   PCmd_IntlkTripSuppress : ALIAS FOR IntlkTrip.PCmd_Suppress;   // Program Command to Suppress Interlock Trip Alarm
   PCmd_IntlkTripUnsuppress : ALIAS FOR IntlkTrip.PCmd_Unsuppress;   // Program Command to Unsuppress Interlock Trip Alarm
   PCmd_IntlkTripUnshelve : ALIAS FOR IntlkTrip.PCmd_Unshelve;   // Program Command to Unshelve Interlock Trip Alarm
   PCmd_IOFaultAck : ALIAS FOR IOFault.PCmd_Ack;   // Program Command to Acknowledge I/O Fault Alarm
   PCmd_IOFaultSuppress : ALIAS FOR IOFault.PCmd_Suppress;   // Program Command to Suppress I/O Fault Alarm
   PCmd_IOFaultUnsuppress : ALIAS FOR IOFault.PCmd_Unsuppress;   // Program Command to Unsuppress I/O Fault Alarm
   PCmd_IOFaultUnshelve : ALIAS FOR IOFault.PCmd_Unshelve;   // Program Command to Unshelve I/O Fault Alarm
   OCmd_Start : BOOL;   // Operator Command to Start Motor
   OCmd_Stop : BOOL;   // Operator Command to Stop Motor
   OCmd_Bypass : BOOL;   // Operator Command to Bypass all Bypassable Interlocks and Permissives
   OCmd_Check : BOOL;   // Operator Command to Check (not bypass) all Interlocks and Permissives
   MCmd_Disable : BOOL;   // Maintenance Command to Disable Motor
   MCmd_Enable : BOOL;   // Maintenance Command to Enable (allow to run) Motor
   OCmd_AcqLock : ALIAS FOR Mode.OCmd_AcqLock;
   OCmd_Unlock : ALIAS FOR Mode.OCmd_UnlockRel;
   OCmd_Reset : BOOL;   // Operator Command to Reset all Alarms requiring Reset
   OCmd_ResetAckAll : BOOL;   // Operator Command to Reset all Alarms and latched Shed conditions
END_VAR
VAR_OUTPUT
   Out_Run : BOOL; {access Read Only, visible}   // 1=Run Motor, 0=Stop Motor
   Out_Start : BOOL; {access Read Only, visible}   // 1=Start Motor, 0=Motor left in current state
   Out_Stop : BOOL; {access Read Only, visible}   // 1=Stop Motor, 0=Motor left in current state
   Val_Cmd : SINT; {access Read Only}   // Device Command 0=None, 1=Stop, 2=Start
   Val_Fdbk : SINT; {access Read Only}   // Device Feedback 0=Stopped, 1=Running
   Val_Sts : SINT; {access Read Only}   // Device Confirmed Sts 0=? 1=Stopped, 2=Running, 7=Stopping, 8=Starting, 33=Disabled
   Val_Fault : SINT; {access Read Only}   // Device Fault Status 0=None, 16=Fail to Start, 17 = Fail to Stop, 32=I/O Fault, 34=Config Error
   Val_Mode : ALIAS FOR Mode.Val; {access Read Only}
   Val_Owner : DINT; {access Read Only}   // Current Object Owner ID (0=not owned)
   Val_Notify : SINT; {access Read Only}   // Current Alarm Level and Acknowledgement (enumeration)
   Sts_Stopped : BOOL := 1; {access Read Only, visible}   // 1=Motor requested to stop and is confirmed stopped
   Sts_Starting : BOOL; {access Read Only, visible}   // 1=Motor requested to run and awaiting run feedback
   Sts_Running : BOOL; {access Read Only, visible}   // 1=Motor requested to run and is confirmed running
   Sts_Stopping : BOOL; {access Read Only, visible}   // 1=Motor requested to stop and awaiting stopped feedback
   Sts_Available : BOOL; {access Read Only}   // 1=Motor available for control by automation (Prog)
   Sts_Bypass : BOOL; {access Read Only}   // 1=Bypassable Interlocks and Permissives are Bypassed
   Sts_BypActive : BOOL; {access Read Only}   // 1=Bypassing Active (Bypassed or Maintenance)
   Sts_Disabled : BOOL; {access Read Only}   // 1=Motor is Disabled
   Sts_NotRdy : BOOL; {access Read Only}   // 1=Motor is Not Ready to Run (independent of Mode)
   Sts_MaintByp : BOOL; {access Read Only}   // 1=A Maintenance Bypass is Active, display icon
   Sts_AlmInh : BOOL; {access Read Only}   // 1=An Alarm is Shelved, Disabled or Suppressed: display icon
   Sts_Err : BOOL; {access Read Only, visible}   // 1=Error in Config: see detail bits for reason
   Err_Timer : BOOL; {access Read Only}   // 1=Error in Config: Start/Stop Check timer preset (use 0 to 2147483)
   Err_Sim : BOOL; {access Read Only}   // 1=Error in Config: Simulation timer preset (use 0 to 2147483)
   Err_Alarm : BOOL; {access Read Only}   // 1=Error in Config: Alarm Min On Time, Shelf Time, Severity
   Sts_Hand : ALIAS FOR Mode.Sts_Hand; {access Read Only, visible}
   Sts_Maint : ALIAS FOR Mode.Sts_Maint; {access Read Only, visible}
   Sts_Ovrd : ALIAS FOR Mode.Sts_Ovrd; {access Read Only, visible}
   Sts_Prog : ALIAS FOR Mode.Sts_Prog; {access Read Only, visible}
   Sts_Oper : ALIAS FOR Mode.Sts_Oper; {access Read Only, visible}
   Sts_ProgOperLock : ALIAS FOR Mode.Sts_ProgOperLock; {access Read Only}
   Sts_NoMode : ALIAS FOR Mode.Sts_NoMode; {access Read Only}
   Sts_FailToStart : ALIAS FOR FailToStart.Inp;   // 1=Motor Failed to Start (one-shot)
   Alm_FailToStart : ALIAS FOR FailToStart.Alm;   // 1=Motor Fail to Start Alarm
   Ack_FailToStart : ALIAS FOR FailToStart.Ack;   // 1=Fail to Start Alarm has been acknowledged
   Sts_FailToStartDisabled : ALIAS FOR FailToStart.Disabled;   // 1=Fail to Start Alarm has been Disabled by Maintenance
   Sts_FailToStartShelved : ALIAS FOR FailToStart.Shelved;   // 1=Fail to Start Alarm has been Shelved by Operator
   Sts_FailToStartSuppressed : ALIAS FOR FailToStart.Suppressed;   // 1=Fail to Start Alarm has been Suppressed by Program
   Sts_FailToStop : ALIAS FOR FailToStop.Inp;   // 1=Motor Failed to Stop
   Alm_FailToStop : ALIAS FOR FailToStop.Alm;   // 1=Motor Fail to Stop Alarm
   Ack_FailToStop : ALIAS FOR FailToStop.Ack;   // 1=Fail to Stop Alarm has been acknowledged
   Sts_FailToStopDisabled : ALIAS FOR FailToStop.Disabled;   // 1=Fail to Stop Alarm has been Disabled by Maintenance
   Sts_FailToStopShelved : ALIAS FOR FailToStop.Shelved;   // 1=Fail to Stop Alarm has been Shelved by Operator
   Sts_FailToStopSuppressed : ALIAS FOR FailToStop.Suppressed;   // 1=Fail to Stop Alarm has been Suppressed by Program
   Sts_IntlkTrip : ALIAS FOR IntlkTrip.Inp;   // 1=Motor stopped by an Interlock NOT OK (one-shot)
   Alm_IntlkTrip : ALIAS FOR IntlkTrip.Alm;   // 1=Alarm: Motor stopped by an Interlock NOT OK
   Ack_IntlkTrip : ALIAS FOR IntlkTrip.Ack;   // 1=Interlock Trip Alarm has been acknowledged
   Sts_IntlkTripDisabled : ALIAS FOR IntlkTrip.Disabled;   // 1=Interlock Trip Alarm has been Disabled by Maintenance
   Sts_IntlkTripShelved : ALIAS FOR IntlkTrip.Shelved;   // 1=Interlock Trip Alarm has been Shelved by Operator
   Sts_IntlkTripSuppressed : ALIAS FOR IntlkTrip.Suppressed;   // 1=Interlock Trip Alarm has been Suppressed by Program
   Sts_IOFault : ALIAS FOR IOFault.Inp;   // I/O Comm Fault Status (0=OK, 1=Bad)
   Alm_IOFault : ALIAS FOR IOFault.Alm;   // 1=I/O Fault Alarm
   Ack_IOFault : ALIAS FOR IOFault.Ack;   // 1=I/O Fault Alarm has been acknowledged
   Sts_IOFaultDisabled : ALIAS FOR IOFault.Disabled;   // 1=I/O Fault Alarm has been Disabled by Maintenance
   Sts_IOFaultShelved : ALIAS FOR IOFault.Shelved;   // 1=I/O Fault Alarm has been Shelved by Operator
   Sts_IOFaultSuppressed : ALIAS FOR IOFault.Suppressed;   // 1=I/O Fault Alarm has been Suppressed by Program
   Rdy_Start : BOOL; {access Read Only}   // 1=Ready to receive OCmd_Start (enables HMI button)
   Rdy_Stop : BOOL; {access Read Only}   // 1=Ready to receive OCmd_Stop (enables HMI button)
   Rdy_Bypass : BOOL; {access Read Only}   // 1=Ready to receive OCmd_Bypass (enables HMI button)
   Rdy_Check : BOOL; {access Read Only}   // 1=Ready to receive OCmd_Check (enables HMI button)
   Rdy_Disable : BOOL; {access Read Only}   // 1=Ready to receive MCmd_Disable (enables HMI button)
   Rdy_Enable : BOOL; {access Read Only}   // 1=Ready to receive MCmd_Enable (enables HMI button)
   Rdy_Reset : BOOL; {access Read Only}   // 1=At least one Alarm or Latched Shed requires Reset
   Rdy_ResetAckAll : BOOL; {access Read Only}   // 1=At least one Alarm or latched Shed condition requires Reset or Ack
   P_Motor : BOOL;   // Unique Parameter Name for auto - discovery
END_VAR
VAR
   Mode : P_Mode := (Cfg_PCmdClear := 1, Cfg_OvrdOverLock := 1, Sts_Oper := 1);   // Motor Mode Selection
   IOFault : P_Alarm := (Inp := 1, Cfg_Exists := 1, Cfg_AckReqd := 1, Cfg_AllowDisable := 1, Cfg_PCmdClear := 1, Cfg_Severity := 3, Cfg_AlmMinOnT := 5, Cfg_MaxShelfT := 480, PCfg_AllowExist := 1, Ack := 1);   // I/O Fault Alarm
   IntlkTrip : P_Alarm := (Inp := 1, Cfg_Exists := 1, Cfg_AckReqd := 1, Cfg_AllowShelve := 1, Cfg_AllowDisable := 1, Cfg_PCmdClear := 1, Cfg_Severity := 3, Cfg_AlmMinOnT := 5, Cfg_MaxShelfT := 480, PCfg_AllowExist := 1, Ack := 1);   // Interlock Trip Alarm
   FailToStop : P_Alarm := (Inp := 1, Cfg_Exists := 1, Cfg_AckReqd := 1, Cfg_AllowDisable := 1, Cfg_PCmdClear := 1, Cfg_Severity := 3, Cfg_AlmMinOnT := 5, Cfg_MaxShelfT := 480, PCfg_AllowExist := 1, Ack := 1);   // Motor Failed to Stop Alarm
   FailToStart : P_Alarm := (Inp := 1, Cfg_Exists := 1, Cfg_AckReqd := 1, Cfg_AllowDisable := 1, Cfg_PCmdClear := 1, Cfg_Severity := 3, Cfg_AlmMinOnT := 5, Cfg_MaxShelfT := 480, PCfg_AllowExist := 1, Ack := 1);   // Motor Failed to Start Alarm
   Cfg_Tag : STRING_20 := 'P_Motor';   // Tagname for display on HMI
   Cfg_Label : STRING_20 := 'P_Motor';   // Label for graphic symbol displayed on HMI
   Cfg_Desc : STRING_40 := 'InFeed Pump';   // Description for display on HMI
   Wrk_Run : BOOL; {access None}   // 1=Motor should be "running", 0=should be "stopped"
   Wrk_SimRunT : TIMER; {access None}   // Simulation Delay until Running
   Wrk_StopT : TIMER; {access None}   // Stop Check Timer
   Wrk_StartT : TIMER; {access None}   // Start Check Timer
   Wrk_SimStopT : TIMER; {access None}   // Simulation Delay until Stopped
   Wrk_RunFdbk : BOOL; {access None}   // Run Feedback based on mode, simulation, etc. 1=running
   Wrk_Notify : DINT; {access None}   // Buffer for building Val_Notify
   Wrk_Bypass : BOOL; {access None}   // Internal Bypassable Permissives and Interlocks are Bypassed flag
   Wrk_Disabled : BOOL; {access None}   // Internal Motor is Disabled
   Inf_Tab : SINT;   // Tab to display (FTView ME)
   Wrk_Cmd : SINT; {access None}   // Buffer for building Val_Cmd
   Wrk_Sts : SINT; {access None}   // Buffer for building Val_Sts
   Wrk_Fault : SINT; {access None}   // Buffer for building Val_Fault
   Wrk_Retrigger : BOOL; {access None}   // Maint Start issued while running or Stop while stopped
   Wrk_FailToStart : BOOL; {access None}   // Fail to Start Fault (latched) stops motor and requires reset
   Wrk_IOFault : BOOL; {access None}   // I/O Fault (latched) stops motor and requires reset
   Inf_Type : STRING_16_UDT := 'P_Motor'; {access Read Only}   // Type identifier for HMI navigation
   Inf_Lib : STRING_12 := 'RA-BAS'; {access Read Only}   // Display Library for Faceplate call-up
END_VAR

ROUTINE EnableInFalse   (* ladder *)
// Disabled is asserted; Outputs OFF; Run Status shown but Alarms disabled
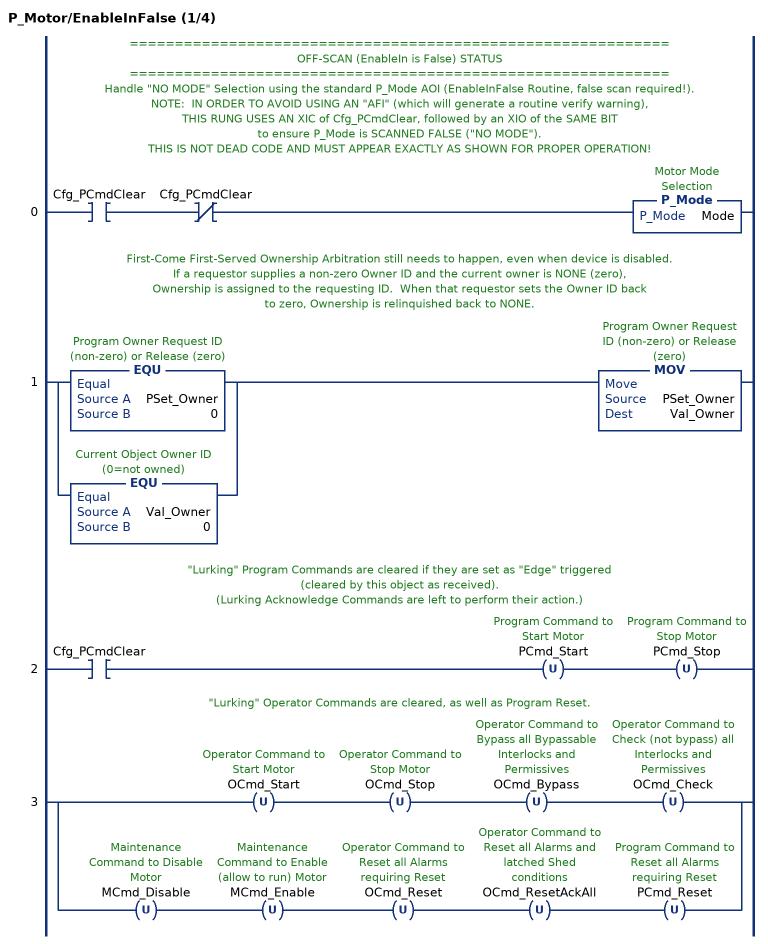
   // ============================================================
   // OFF-SCAN (EnableIn is False) STATUS
   // ============================================================
   // Handle "NO MODE" Selection using the standard P_Mode AOI (EnableInFalse Routine, false scan required!).
   // NOTE:  IN ORDER TO AVOID USING AN "AFI" (which will generate a routine verify warning),
   // THIS RUNG USES AN XIC of Cfg_PCmdClear, followed by an XIO of the SAME BIT
   // to ensure P_Mode is SCANNED FALSE ("NO MODE").
   // THIS IS NOT DEAD CODE AND MUST APPEAR EXACTLY AS SHOWN FOR PROPER OPERATION!
   0: XIC(Cfg_PCmdClear)XIO(Cfg_PCmdClear)P_Mode(Mode);
   // First-Come First-Served Ownership Arbitration still needs to happen, even when device is disabled.
   // If a requestor supplies a non-zero Owner ID and the current owner is NONE (zero),
   // Ownership is assigned to the requesting ID.  When that requestor sets the Owner ID back
   // to zero, Ownership is relinquished back to NONE.
   1: [EQU(PSet_Owner,0) ,EQU(Val_Owner,0) ]MOV(PSet_Owner,Val_Owner);
   // "Lurking" Program Commands are cleared if they are set as "Edge" triggered
   // (cleared by this object as received).
   // (Lurking Acknowledge Commands are left to perform their action.)
   2: XIC(Cfg_PCmdClear)OTU(PCmd_Start)OTU(PCmd_Stop);
   // "Lurking" Operator Commands are cleared, as well as Program Reset.
   3: [OTU(OCmd_Start) OTU(OCmd_Stop) OTU(OCmd_Bypass) OTU(OCmd_Check) ,OTU(MCmd_Disable) OTU(MCmd_Enable) OTU(OCmd_Reset) OTU(OCmd_ResetAckAll) OTU(PCmd_Reset) ];
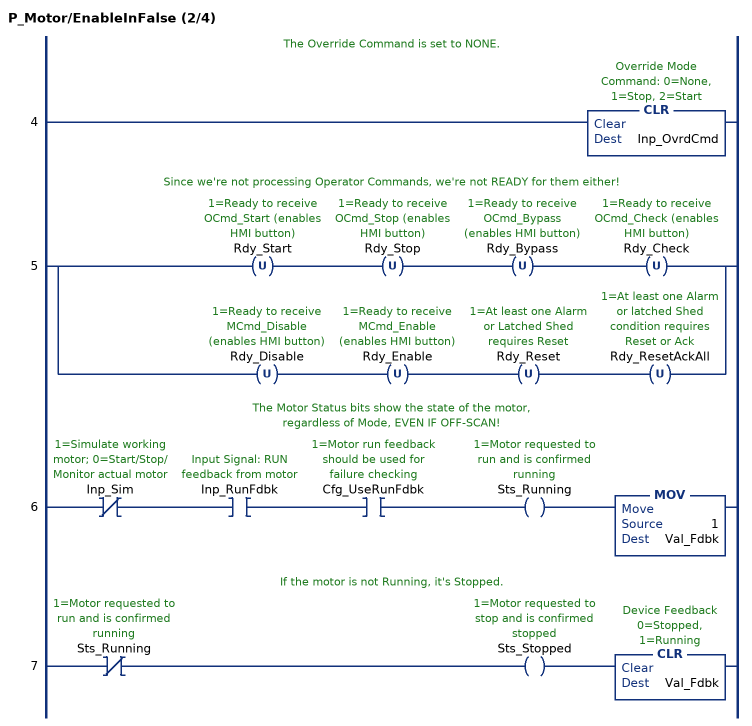
   // The Override Command is set to NONE.
   4: CLR(Inp_OvrdCmd);
   // Since we're not processing Operator Commands, we're not READY for them either!
   5: [OTU(Rdy_Start) OTU(Rdy_Stop) OTU(Rdy_Bypass) OTU(Rdy_Check) ,OTU(Rdy_Disable) OTU(Rdy_Enable) OTU(Rdy_Reset) OTU(Rdy_ResetAckAll) ];
   // The Motor Status bits show the state of the motor,
   // regardless of Mode, EVEN IF OFF-SCAN!
   6: XIO(Inp_Sim)XIC(Inp_RunFdbk)XIC(Cfg_UseRunFdbk)OTE(Sts_Running)MOV(1,Val_Fdbk);
   // If the motor is not Running, it's Stopped.
   7: XIO(Sts_Running)OTE(Sts_Stopped)CLR(Val_Fdbk);
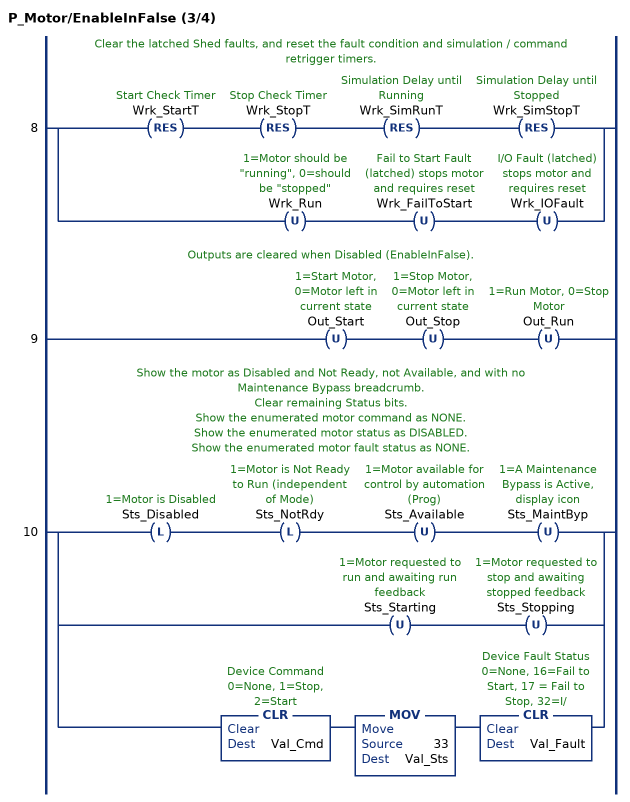
   // Clear the latched Shed faults, and reset the fault condition and simulation / command retrigger timers.
   8: [RES(Wrk_StartT) RES(Wrk_StopT) RES(Wrk_SimRunT) RES(Wrk_SimStopT) ,OTU(Wrk_Run) OTU(Wrk_FailToStart) OTU(Wrk_IOFault) ];
   // Outputs are cleared when Disabled (EnableInFalse).
   9: OTU(Out_Start)OTU(Out_Stop)OTU(Out_Run);
   // Show the motor as Disabled and Not Ready, not Available, and with no
   // Maintenance Bypass breadcrumb.
   // Clear remaining Status bits.
   // Show the enumerated motor command as NONE.
   // Show the enumerated motor status as DISABLED.
   // Show the enumerated motor fault status as NONE.
   10: [OTL(Sts_Disabled) OTL(Sts_NotRdy) OTU(Sts_Available) OTU(Sts_MaintByp) ,OTU(Sts_Starting) OTU(Sts_Stopping) ,CLR(Val_Cmd) MOV(33,Val_Sts) CLR(Val_Fault) ];
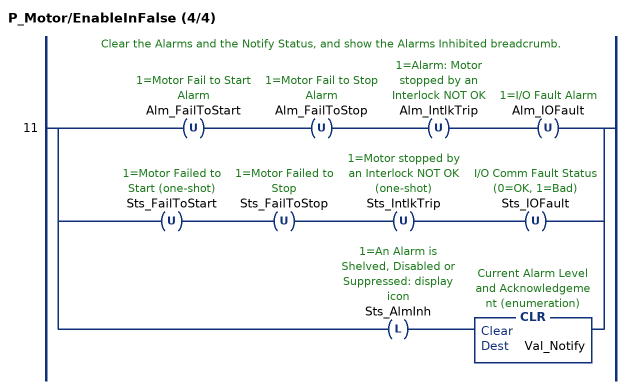
   // Clear the Alarms and the Notify Status, and show the Alarms Inhibited breadcrumb.
   11: [OTU(Alm_FailToStart) OTU(Alm_FailToStop) OTU(Alm_IntlkTrip) OTU(Alm_IOFault) ,OTU(Sts_FailToStart) OTU(Sts_FailToStop) OTU(Sts_IntlkTrip) OTU(Sts_IOFault) ,OTL(Sts_AlmInh) CLR(Val_Notify) ];
END_ROUTINE

ROUTINE Logic   (* ladder *)
// Normal Scan: control / monitor single speed motor
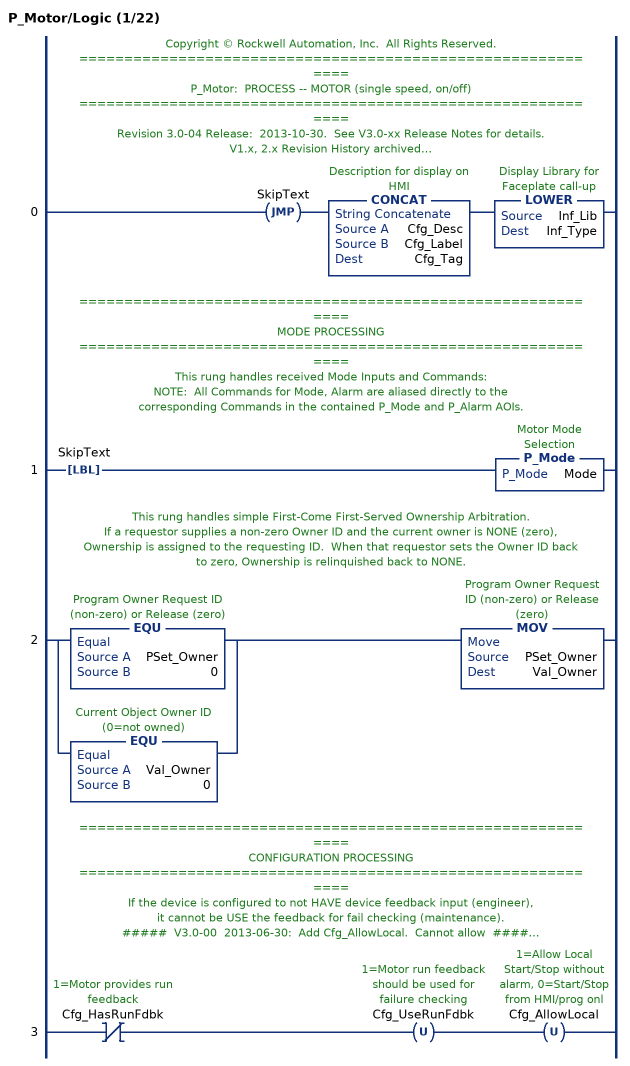
   // Copyright © Rockwell Automation, Inc.  All Rights Reserved.
   // ============================================================
   // P_Motor:  PROCESS -- MOTOR (single speed, on/off)
   // ============================================================
   // Revision 3.0-04 Release:  2013-10-30.  See V3.0-xx Release Notes for details.
   // V1.x, 2.x Revision History archived.
   // V3.0-00:  2013-06-30.  Added Inf_Lib.  Added Cfg_AllowLocal, Cfg_OperStopPrio,
   // Cfg_HasOvldObj.  Using P_Alarm 3.0, P_Mode 3.0.
   // V3.0-01:  2013-07-30.  Modified Parameter descriptions only.
   // V3.0-02:  2013-09-03.  Modified to ensure Out_Stop always pulses
   // whenever a stop command is received, regardless of run
   // feedback state.  Modified Parameter descriptions.
   // V3.0-03:  2013-09-10.  Corrected modification above for operation
   // in simulation and for all start, stop and not-ready conditions.
   // V3.0-04:  2013-10-30.  Corrected Parameter descriptions and default
   // configuration values for alarms only.
   // Modified default Parameter values.
   // ============================================================
   // This Instruction controls and monitors a single-speed motor
   // (FVNR, soft-start, etc.) and provides:
   // *  Monitoring of run feedback, display of actual motor status
   // *  Detection of Failure to Start, Failure to Stop
   // *  Monitoring of a Permissive condition to allow starting
   // * Monitoring of an Interlock condition to stop / prevent starting
   // * Simulation, providing feedback of a working motor while disabling outputs
   // * Monitoring of I/O communication faults
   // * Alarms for Fail to Start, Fail to Stop, Interlock Trip, I/O Fault
   // * Options to shed (stop motor) on Fail to Start or I/O Fault
   // * Option to automatically reset faults and alarms when operator commands
   // motor to start or stop
   // * Supports HMI "breadcrumbs" for Alarm Inhibited, Bad Configuration,
   // Not Ready, Maintenance Bypass Active
   // * "Available" status for use by automation logic to know whether motor
   // can be controlled by other objects.
   // Modes are provided by a P_Mode AOI instance.
   // Alarms are provided by P_Alarm AOI instances.
   // Modes of operation: Operator, Program, Override, Maintenance, Hand
   // ============================================================
   // SHOW LOCAL STRINGS
   // ============================================================
   // The STRINGs containing the text associated with each instance of this
   // instruction cannot be Input or Output Parameters, because STRINGs are not
   //  'atomic' types. (Inputs and Outputs must be SINT, INT, DINT, REAL, or BOOL.)
   // In order to make it easier to find and configure these STRINGs, this rung
   // was added.  THE JMP (and the LBL on the following rung)
   // MUST NOT BE REMOVED!!!
   // To view the STRINGs, go to the instruction instance (in LD or FBD), RIGHT-click
   // to bring up the context menu and select "Open Instruction Logic".
   // This rung will appear with the STRING values for the selected instance.
   // You may double-click the STRING values here to modify them as well.
   0: JMP(SkipText)CONCAT(Cfg_Desc,Cfg_Label,Cfg_Tag)LOWER(Inf_Lib,Inf_Type);
   // ============================================================
   // MODE PROCESSING
   // ============================================================
   // This rung handles received Mode Inputs and Commands:
   // NOTE:  All Commands for Mode, Alarm are aliased directly to the
   // corresponding Commands in the contained P_Mode and P_Alarm AOIs.
   1: LBL(SkipText)P_Mode(Mode);
   // This rung handles simple First-Come First-Served Ownership Arbitration.
   // If a requestor supplies a non-zero Owner ID and the current owner is NONE (zero),
   // Ownership is assigned to the requesting ID.  When that requestor sets the Owner ID back
   // to zero, Ownership is relinquished back to NONE.
   2: [EQU(PSet_Owner,0) ,EQU(Val_Owner,0) ]MOV(PSet_Owner,Val_Owner);
   // ============================================================
   // CONFIGURATION PROCESSING
   // ============================================================
   // If the device is configured to not HAVE device feedback input (engineer),
   // it cannot be USE the feedback for fail checking (maintenance).
   // #####  V3.0-00  2013-06-30:  Add Cfg_AllowLocal.  Cannot allow  #####
   // #####  local start/stop  if run feedback does not exist to monitor for it.  #####
   3: XIO(Cfg_HasRunFdbk)OTU(Cfg_UseRunFdbk)OTU(Cfg_AllowLocal);
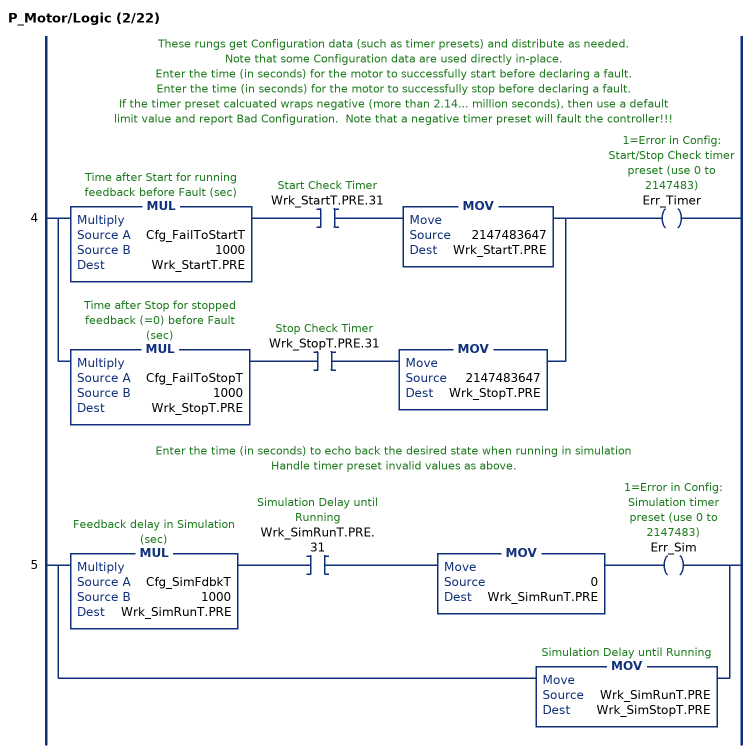
   // These rungs get Configuration data (such as timer presets) and distribute as needed.
   // Note that some Configuration data are used directly in-place.
   // Enter the time (in seconds) for the motor to successfully start before declaring a fault.
   // Enter the time (in seconds) for the motor to successfully stop before declaring a fault.
   // If the timer preset calcuated wraps negative (more than 2.14... million seconds), then use a default
   // limit value and report Bad Configuration.  Note that a negative timer preset will fault the controller!!!
   4: [MUL(Cfg_FailToStartT,1000,Wrk_StartT.PRE) XIC(Wrk_StartT.PRE.31) MOV(2147483647,Wrk_StartT.PRE) ,MUL(Cfg_FailToStopT,1000,Wrk_StopT.PRE) XIC(Wrk_StopT.PRE.31) MOV(2147483647,Wrk_StopT.PRE) ]OTE(Err_Timer);
   // Enter the time (in seconds) to echo back the desired state when running in simulation
   // Handle timer preset invalid values as above.
   5: [MUL(Cfg_SimFdbkT,1000,Wrk_SimRunT.PRE) XIC(Wrk_SimRunT.PRE.31) MOV(0,Wrk_SimRunT.PRE) OTE(Err_Sim) ,MOV(Wrk_SimRunT.PRE,Wrk_SimStopT.PRE) ];
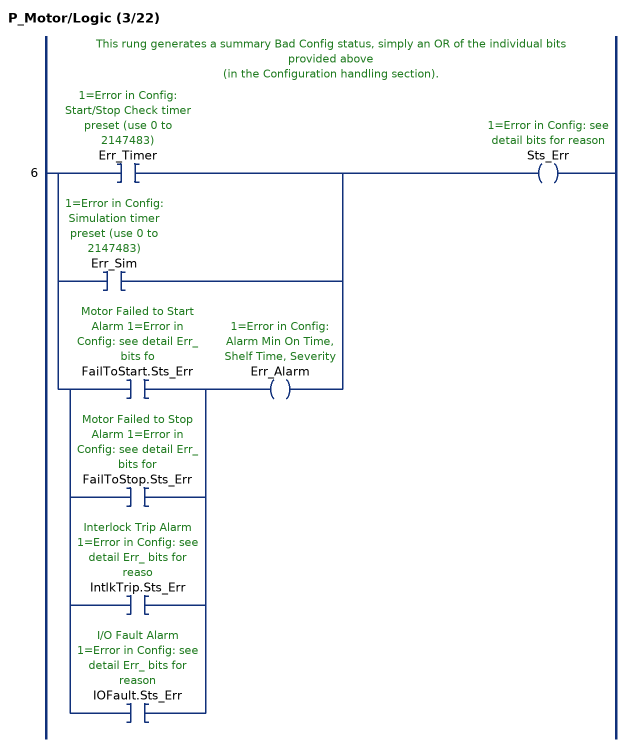
   // This rung generates a summary Bad Config status, simply an OR of the individual bits provided above
   // (in the Configuration handling section).
   6: [XIC(Err_Timer) ,XIC(Err_Sim) ,[XIC(FailToStart.Sts_Err) ,XIC(FailToStop.Sts_Err) ,XIC(IntlkTrip.Sts_Err) ,XIC(IOFault.Sts_Err) ] OTE(Err_Alarm) ]OTE(Sts_Err);
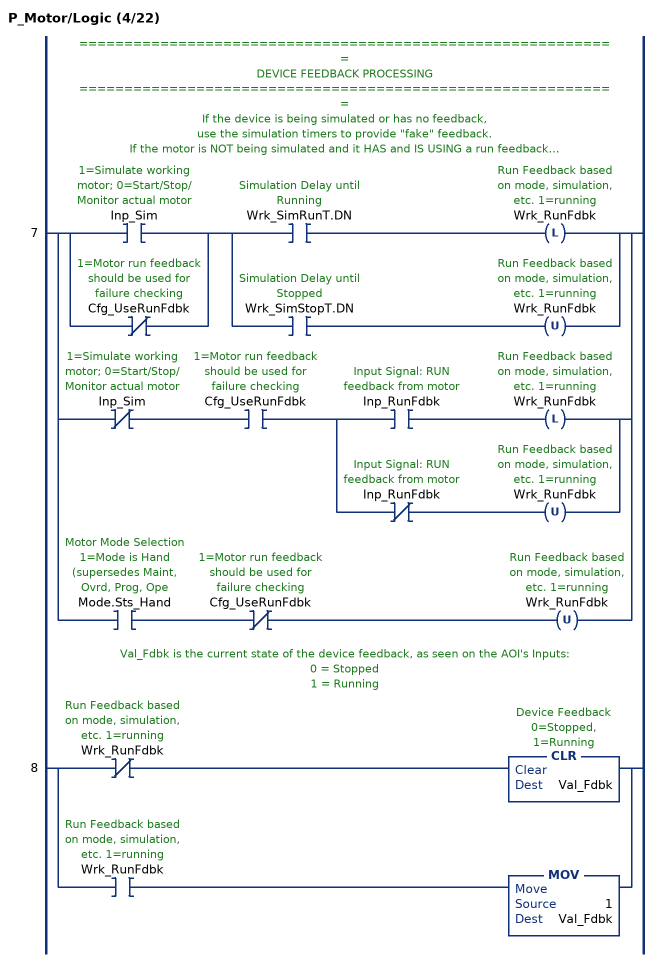
   // ============================================================
   // DEVICE FEEDBACK PROCESSING
   // ============================================================
   // If the device is being simulated or has no feedback,
   // use the simulation timers to provide "fake" feedback.
   // If the motor is NOT being simulated and it HAS and IS USING a run feedback,
   // use the state of the run feedback input as the motor run state.
   7: [[XIC(Inp_Sim) ,XIO(Cfg_UseRunFdbk) ] [XIC(Wrk_SimRunT.DN) OTL(Wrk_RunFdbk) ,XIC(Wrk_SimStopT.DN) OTU(Wrk_RunFdbk) ] ,XIO(Inp_Sim) XIC(Cfg_UseRunFdbk) [XIC(Inp_RunFdbk) OTL(Wrk_RunFdbk) ,XIO(Inp_RunFdbk) OTU(Wrk_RunFdbk) ] ,XIC(Mode.Sts_Hand) XIO(Cfg_UseRunFdbk) OTU(Wrk_RunFdbk) ];
   // Val_Fdbk is the current state of the device feedback, as seen on the AOI's Inputs:
   // 0 = Stopped
   // 1 = Running
   8: [XIO(Wrk_RunFdbk) CLR(Val_Fdbk) ,XIC(Wrk_RunFdbk) MOV(1,Val_Fdbk) ];
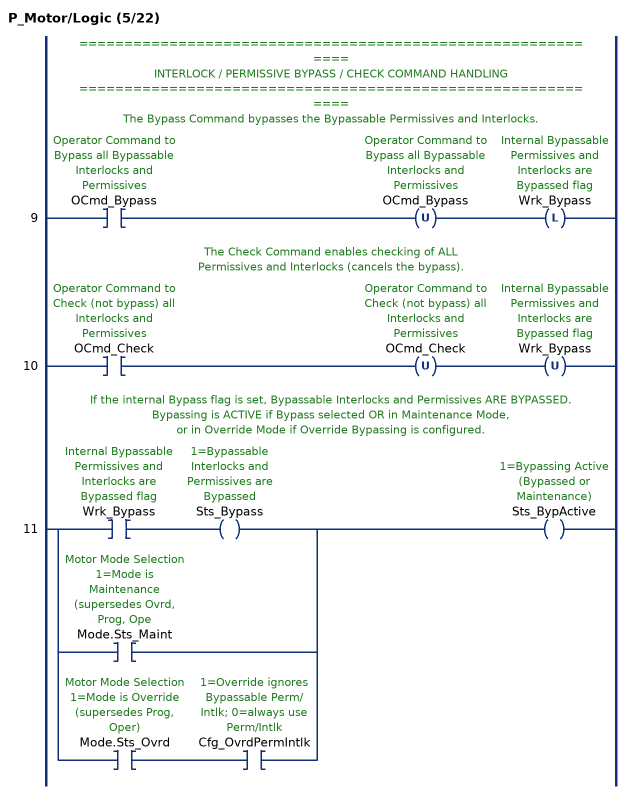
   // ============================================================
   // INTERLOCK / PERMISSIVE BYPASS / CHECK COMMAND HANDLING
   // ============================================================
   // The Bypass Command bypasses the Bypassable Permissives and Interlocks.
   9: XIC(OCmd_Bypass)OTU(OCmd_Bypass)OTL(Wrk_Bypass);
   // The Check Command enables checking of ALL
   // Permissives and Interlocks (cancels the bypass).
   10: XIC(OCmd_Check)OTU(OCmd_Check)OTU(Wrk_Bypass);
   // If the internal Bypass flag is set, Bypassable Interlocks and Permissives ARE BYPASSED.
   // Bypassing is ACTIVE if Bypass selected OR in Maintenance Mode,
   // or in Override Mode if Override Bypassing is configured.
   11: [XIC(Wrk_Bypass) OTE(Sts_Bypass) ,XIC(Mode.Sts_Maint) ,XIC(Mode.Sts_Ovrd) XIC(Cfg_OvrdPermIntlk) ]OTE(Sts_BypActive);
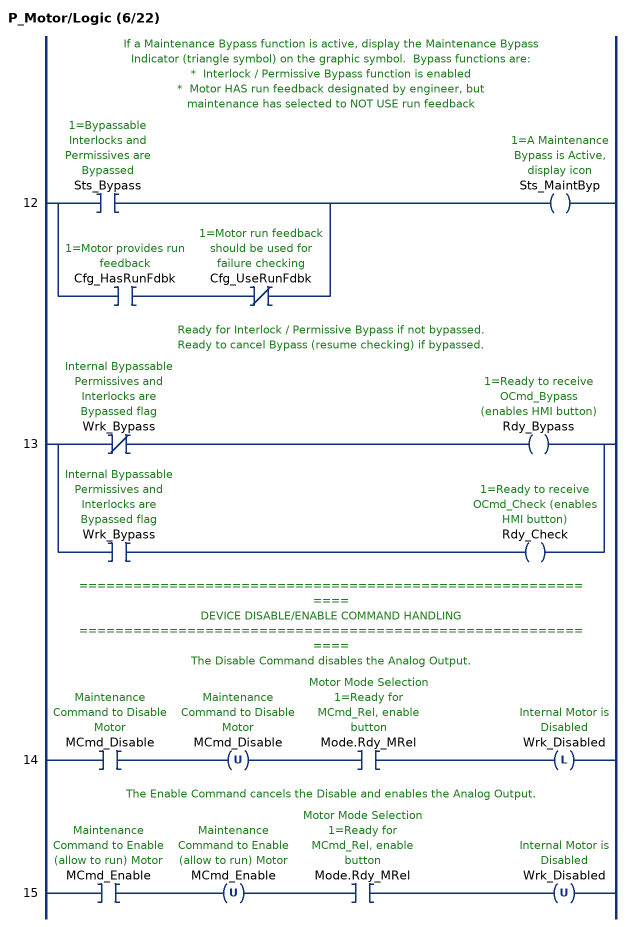
   // If a Maintenance Bypass function is active, display the Maintenance Bypass
   // Indicator (triangle symbol) on the graphic symbol.  Bypass functions are:
   // *  Interlock / Permissive Bypass function is enabled
   // *  Motor HAS run feedback designated by engineer, but
   // maintenance has selected to NOT USE run feedback
   12: [XIC(Sts_Bypass) ,XIC(Cfg_HasRunFdbk) XIO(Cfg_UseRunFdbk) ]OTE(Sts_MaintByp);
   // Ready for Interlock / Permissive Bypass if not bypassed.
   // Ready to cancel Bypass (resume checking) if bypassed.
   13: [XIO(Wrk_Bypass) OTE(Rdy_Bypass) ,XIC(Wrk_Bypass) OTE(Rdy_Check) ];
   // ============================================================
   // DEVICE DISABLE/ENABLE COMMAND HANDLING
   // ============================================================
   // The Disable Command disables the Analog Output.
   14: XIC(MCmd_Disable)OTU(MCmd_Disable)XIC(Mode.Rdy_MRel)OTL(Wrk_Disabled);
   // The Enable Command cancels the Disable and enables the Analog Output.
   15: XIC(MCmd_Enable)OTU(MCmd_Enable)XIC(Mode.Rdy_MRel)OTU(Wrk_Disabled);
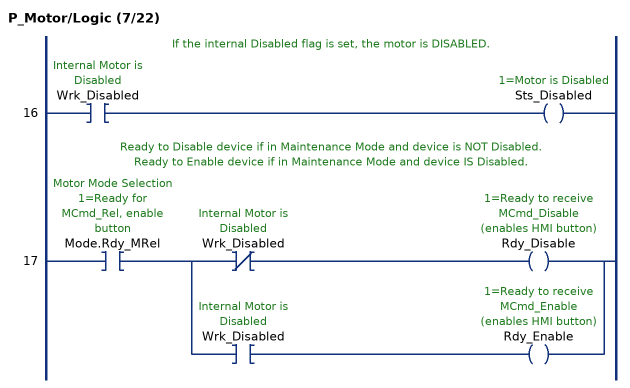
   // If the internal Disabled flag is set, the motor is DISABLED.
   16: XIC(Wrk_Disabled)OTE(Sts_Disabled);
   // Ready to Disable device if in Maintenance Mode and device is NOT Disabled.
   // Ready to Enable device if in Maintenance Mode and device IS Disabled.
   17: XIC(Mode.Rdy_MRel)[XIO(Wrk_Disabled) OTE(Rdy_Disable) ,XIC(Wrk_Disabled) OTE(Rdy_Enable) ];
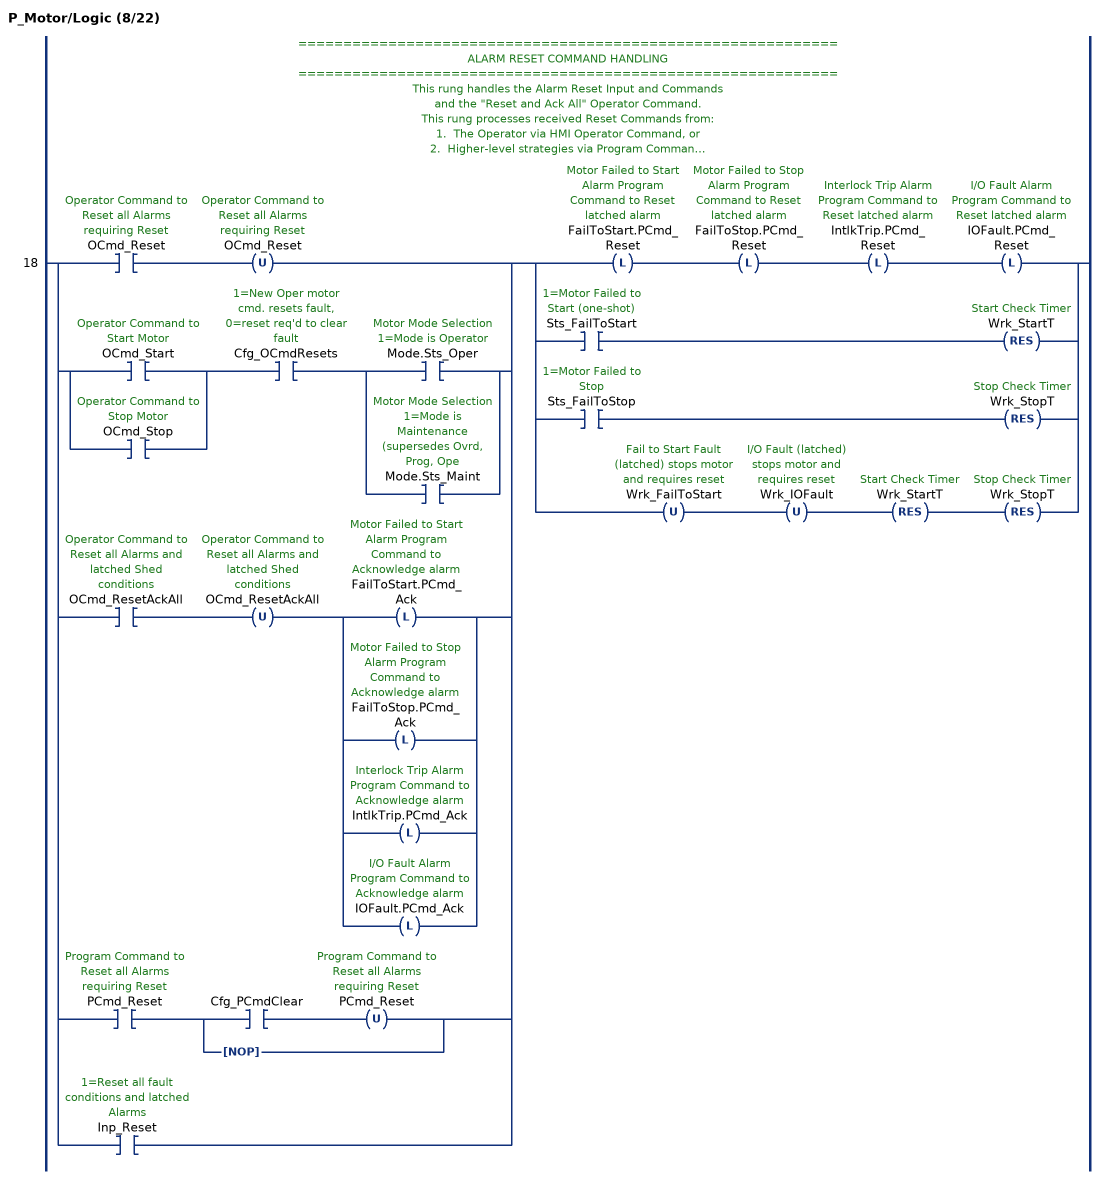
   // ============================================================
   // ALARM RESET COMMAND HANDLING
   // ============================================================
   // This rung handles the Alarm Reset Input and Commands
   // and the "Reset and Ack All" Operator Command.
   // This rung processes received Reset Commands from:
   // 1.  The Operator via HMI Operator Command, or
   // 2.  Higher-level strategies via Program Command
   // 3.  Pushbuttons or other block via Input
   // 4.  Resets initiated by other device Operator Commands (if configured to do so)
   // and forwards the Reset to ALL Alarms and latched Shed conditions.
   18: [[XIC(OCmd_Reset) OTU(OCmd_Reset) ,[XIC(OCmd_Start) ,XIC(OCmd_Stop) ] XIC(Cfg_OCmdResets) [XIC(Mode.Sts_Oper) ,XIC(Mode.Sts_Maint) ] ] ,XIC(OCmd_ResetAckAll) OTU(OCmd_ResetAckAll) [OTL(FailToStart.PCmd_Ack) ,OTL(FailToStop.PCmd_Ack) ,OTL(IntlkTrip.PCmd_Ack) ,OTL(IOFault.PCmd_Ack) ] ,XIC(PCmd_Reset) [XIC(Cfg_PCmdClear) OTU(PCmd_Reset) ,NOP() ] ,XIC(Inp_Reset) ][OTL(FailToStart.PCmd_Reset) OTL(FailToStop.PCmd_Reset) OTL(IntlkTrip.PCmd_Reset) OTL(IOFault.PCmd_Reset) ,XIC(Sts_FailToStart) RES(Wrk_StartT) ,XIC(Sts_FailToStop) RES(Wrk_StopT) ,OTU(Wrk_FailToStart) OTU(Wrk_IOFault) RES(Wrk_StartT) RES(Wrk_StopT) ];
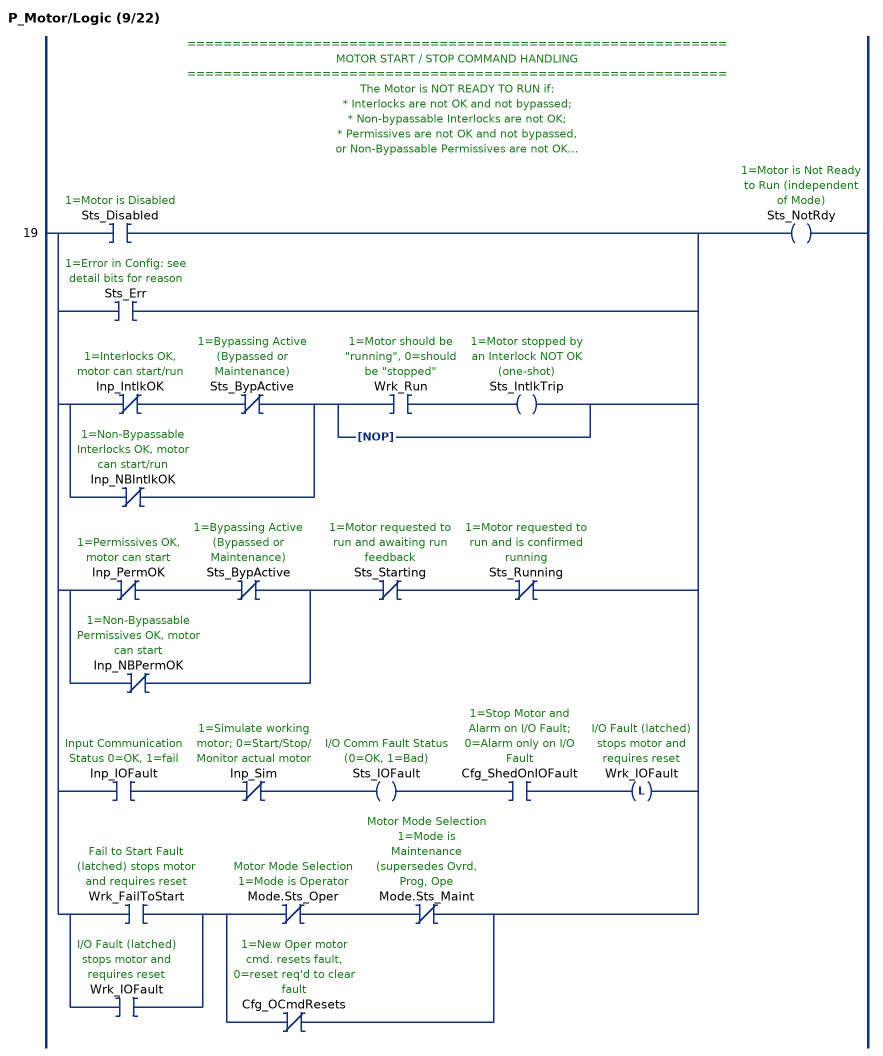
   // ============================================================
   // MOTOR START / STOP COMMAND HANDLING
   // ============================================================
   // The Motor is NOT READY TO RUN if:
   // * Interlocks are not OK and not bypassed;
   // * Non-bypassable Interlocks are not OK;
   // * Permissives are not OK and not bypassed,
   // or Non-Bypassable Permissives are not OK,
   // and the motor is not already starting or running;
   // * There's an I/O failure and the motor is NOT being simulated;
   // * The motor has a Fail to Start or Fail to Stop that has not been reset;
   // * The motor is disabled by Maintenance.
   19: [XIC(Sts_Disabled) ,XIC(Sts_Err) ,[XIO(Inp_IntlkOK) XIO(Sts_BypActive) ,XIO(Inp_NBIntlkOK) ] [XIC(Wrk_Run) OTE(Sts_IntlkTrip) ,NOP() ] ,[XIO(Inp_PermOK) XIO(Sts_BypActive) ,XIO(Inp_NBPermOK) ] XIO(Sts_Starting) XIO(Sts_Running) ,XIC(Inp_IOFault) XIO(Inp_Sim) OTE(Sts_IOFault) XIC(Cfg_ShedOnIOFault) OTL(Wrk_IOFault) ,[XIC(Wrk_FailToStart) ,XIC(Wrk_IOFault) ] [XIO(Mode.Sts_Oper) XIO(Mode.Sts_Maint) ,XIO(Cfg_OCmdResets) ] ]OTE(Sts_NotRdy);
